screen "1002_Process Value Mixing Head" 1280x800, template "Navigation"
   on GenerateScreen: SetBit("DB704_MH_Value_Read")
   Group "Group" at 107,163 size 1065x534
   TextField "Text field_1" at 500,138 size 280x25; Text 'Process values metering unit / Process values mixing head'
   TextField "Text field_2" at 138,222 size 112x25; Text 'Module No.'
   TextField "Text field_3" at 138,256 size 81x25; Text 'Address'
   TextField "Text field_4" at 138,290 size 64x25; Text 'Offset'
   TextField "Text field_5" at 138,323 size 96x25; Text 'Multiplier'
   TextField "Text field_6" at 138,357 size 174x25; Text 'Min. Value Sensor'
   TextField "Text field_7" at 138,391 size 178x25; Text 'Max. Value Sensor'
   TextField "Text field_10" at 445,189 size 141x25; Text 'Pressure Con2'
   TextField "Text field_11" at 589,189 size 141x25; Text 'Pressure Con3'
   IOField "PV_MeteringUnit_ModulNoPressureCon1" at 313,219 size 122x30; Authorization "User administration"; FormatPattern s9999999
      ProcessValue <- "DB604_PV_Mixinghead_Mixinghead{0}_Pressure_Connection{1}_PV_Conf_ActV_ModulNo"
   IOField "I/O field_2" at 313,253 size 122x30; Authorization "User administration"; FormatPattern s9999999
      ProcessValue <- "DB604_PV_Mixinghead_Mixinghead{0}_Pressure_Connection{1}_PV_Conf_ActV_Address"
   IOField "I/O field_3" at 313,287 size 122x30; Authorization "User administration"; FormatPattern s9999999
      ProcessValue <- "DB604_PV_Mixinghead_Mixinghead{0}_Pressure_Connection{1}_PV_Conf_ActV_OffsetSignal"
   IOField "I/O field_4" at 313,321 size 122x30; Authorization "User administration"; FormatPattern s99999.999
      ProcessValue <- "DB604_PV_Mixinghead_Mixinghead{0}_Pressure_Connection{1}_PV_Conf_ActV_Multiplier"
   IOField "I/O field_5" at 313,355 size 122x30; Authorization "User administration"; FormatPattern s99999
      ProcessValue <- "DB604_PV_Mixinghead_Mixinghead{0}_Pressure_Connection{1}_PV_Conf_ActV_MinValueSensor"
   IOField "I/O field_6" at 313,389 size 122x30; Authorization "User administration"; FormatPattern s9999999
      ProcessValue <- "DB604_PV_Mixinghead_Mixinghead{0}_Pressure_Connection{1}_PV_Conf_ActV_MaxValueSensor"
   IOField "I/O field_8" at 454,219 size 122x30; Authorization "User administration"; FormatPattern s9999999
      ProcessValue <- "DB604_PV_Mixinghead_Mixinghead{0}_Pressure_Connection{2}_PV_Conf_ActV_ModulNo"
   IOField "I/O field_9" at 454,253 size 122x30; Authorization "User administration"; FormatPattern s9999999
      ProcessValue <- "DB604_PV_Mixinghead_Mixinghead{0}_Pressure_Connection{2}_PV_Conf_ActV_Address"
   IOField "I/O field_10" at 454,287 size 122x30; Authorization "User administration"; FormatPattern s9999999
      ProcessValue <- "DB604_PV_Mixinghead_Mixinghead{0}_Pressure_Connection{2}_PV_Conf_ActV_OffsetSignal"
   IOField "I/O field_11" at 454,321 size 122x30; Authorization "User administration"; FormatPattern s99999.999
      ProcessValue <- "DB604_PV_Mixinghead_Mixinghead{0}_Pressure_Connection{2}_PV_Conf_ActV_Multiplier"
   IOField "I/O field_12" at 454,355 size 122x30; Authorization "User administration"; FormatPattern s99999
      ProcessValue <- "DB604_PV_Mixinghead_Mixinghead{0}_Pressure_Connection{2}_PV_Conf_ActV_MinValueSensor"
   IOField "I/O field_13" at 454,389 size 122x30; Authorization "User administration"; FormatPattern s9999999
      ProcessValue <- "DB604_PV_Mixinghead_Mixinghead{0}_Pressure_Connection{2}_PV_Conf_ActV_MaxValueSensor"
   IOField "I/O field_14" at 598,219 size 122x30; Authorization "User administration"; FormatPattern s9999999
      ProcessValue <- "DB604_PV_Mixinghead_Mixinghead{0}_Pressure_Connection{3}_PV_Conf_ActV_ModulNo"
   IOField "I/O field_15" at 598,253 size 122x30; Authorization "User administration"; FormatPattern s9999999
      ProcessValue <- "DB604_PV_Mixinghead_Mixinghead{0}_Pressure_Connection{3}_PV_Conf_ActV_Address"
   IOField "I/O field_16" at 598,287 size 122x30; Authorization "User administration"; FormatPattern s9999999
      ProcessValue <- "DB604_PV_Mixinghead_Mixinghead{0}_Pressure_Connection{3}_PV_Conf_ActV_OffsetSignal"
   IOField "I/O field_17" at 598,321 size 122x30; Authorization "User administration"; FormatPattern s99999.999
      ProcessValue <- "DB604_PV_Mixinghead_Mixinghead{0}_Pressure_Connection{3}_PV_Conf_ActV_Multiplier"
   IOField "I/O field_18" at 598,355 size 122x30; Authorization "User administration"; FormatPattern s99999
      ProcessValue <- "DB604_PV_Mixinghead_Mixinghead{0}_Pressure_Connection{3}_PV_Conf_ActV_MinValueSensor"
   IOField "I/O field_19" at 598,389 size 122x30; Authorization "User administration"; FormatPattern s9999999
      ProcessValue <- "DB604_PV_Mixinghead_Mixinghead{0}_Pressure_Connection{3}_PV_Conf_ActV_MaxValueSensor"
   TextField "Text field_16" at 734,189 size 141x25; Text 'Pressure Con4'
   TextField "Text field_17" at 873,189 size 141x25; Text 'Pressure Con5'
   IOField "I/O field_23" at 882,219 size 122x30; Authorization "User administration"; FormatPattern s9999999
      ProcessValue <- "DB604_PV_Mixinghead_Mixinghead{0}_Pressure_Connection{5}_PV_Conf_ActV_ModulNo"
   IOField "I/O field_24" at 882,253 size 122x30; Authorization "User administration"; FormatPattern s9999999
      ProcessValue <- "DB604_PV_Mixinghead_Mixinghead{0}_Pressure_Connection{5}_PV_Conf_ActV_Address"
   IOField "I/O field_25" at 882,287 size 122x30; Authorization "User administration"; FormatPattern s9999999
      ProcessValue <- "DB604_PV_Mixinghead_Mixinghead{0}_Pressure_Connection{5}_PV_Conf_ActV_OffsetSignal"
   IOField "I/O field_26" at 882,321 size 122x30; Authorization "User administration"; FormatPattern s99999.999
      ProcessValue <- "DB604_PV_Mixinghead_Mixinghead{0}_Pressure_Connection{5}_PV_Conf_ActV_Multiplier"
   IOField "I/O field_27" at 882,355 size 122x30; Authorization "User administration"; FormatPattern s99999
      ProcessValue <- "DB604_PV_Mixinghead_Mixinghead{0}_Pressure_Connection{5}_PV_Conf_ActV_MinValueSensor"
   IOField "I/O field_28" at 882,389 size 122x30; Authorization "User administration"; FormatPattern s9999999
      ProcessValue <- "DB604_PV_Mixinghead_Mixinghead{0}_Pressure_Connection{5}_PV_Conf_ActV_MaxValueSensor"
   TextField "Text field_9" at 304,189 size 141x25; Text 'Pressure Con1'
   TextField "Text field_29" at 1014,191 size 141x25; Text 'Pressure Con6'
   IOField "I/O field_35" at 1023,219 size 122x30; Authorization "User administration"; FormatPattern s9999999
      ProcessValue <- "DB604_PV_Mixinghead_Mixinghead{0}_Pressure_Connection{6}_PV_Conf_ActV_ModulNo"
   IOField "I/O field_36" at 1023,253 size 122x30; Authorization "User administration"; FormatPattern s9999999
      ProcessValue <- "DB604_PV_Mixinghead_Mixinghead{0}_Pressure_Connection{6}_PV_Conf_ActV_Address"
   IOField "I/O field_37" at 1023,287 size 122x30; Authorization "User administration"; FormatPattern s9999999
      ProcessValue <- "DB604_PV_Mixinghead_Mixinghead{0}_Pressure_Connection{6}_PV_Conf_ActV_OffsetSignal"
   IOField "I/O field_38" at 1023,321 size 122x30; Authorization "User administration"; FormatPattern s99999.999
      ProcessValue <- "DB604_PV_Mixinghead_Mixinghead{0}_Pressure_Connection{6}_PV_Conf_ActV_Multiplier"
   IOField "I/O field_39" at 1023,355 size 122x30; Authorization "User administration"; FormatPattern s99999
      ProcessValue <- "DB604_PV_Mixinghead_Mixinghead{0}_Pressure_Connection{6}_PV_Conf_ActV_MinValueSensor"
   IOField "I/O field_40" at 1023,389 size 122x30; Authorization "User administration"; FormatPattern s9999999
      ProcessValue <- "DB604_PV_Mixinghead_Mixinghead{0}_Pressure_Connection{6}_PV_Conf_ActV_MaxValueSensor"
   IOField "I/O field_7" at 739,219 size 122x30; Authorization "User administration"; FormatPattern s9999999
      ProcessValue <- "DB604_PV_Mixinghead_Mixinghead{0}_Pressure_Connection{4}_PV_Conf_ActV_ModulNo"
   IOField "I/O field_20" at 739,253 size 122x30; Authorization "User administration"; FormatPattern s9999999
      ProcessValue <- "DB604_PV_Mixinghead_Mixinghead{0}_Pressure_Connection{4}_PV_Conf_ActV_Address"
   IOField "I/O field_21" at 739,287 size 122x30; Authorization "User administration"; FormatPattern s9999999
      ProcessValue <- "DB604_PV_Mixinghead_Mixinghead{0}_Pressure_Connection{4}_PV_Conf_ActV_OffsetSignal"
   IOField "I/O field_22" at 739,321 size 122x30; Authorization "User administration"; FormatPattern s99999.999
      ProcessValue <- "DB604_PV_Mixinghead_Mixinghead{0}_Pressure_Connection{4}_PV_Conf_ActV_Multiplier"
   IOField "I/O field_29" at 739,355 size 122x30; Authorization "User administration"; FormatPattern s99999
      ProcessValue <- "DB604_PV_Mixinghead_Mixinghead{0}_Pressure_Connection{4}_PV_Conf_ActV_MinValueSensor"
   IOField "I/O field_30" at 739,389 size 122x30; Authorization "User administration"; FormatPattern s9999999
      ProcessValue <- "DB604_PV_Mixinghead_Mixinghead{0}_Pressure_Connection{4}_PV_Conf_ActV_MaxValueSensor"
   TextField "Text field_8" at 138,462 size 112x25; Text 'Module No.'
   TextField "Text field_12" at 138,497 size 81x25; Text 'Address'
   TextField "Text field_13" at 138,532 size 64x25; Text 'Offset'
   TextField "Text field_14" at 138,566 size 96x25; Text 'Multiplier'
   TextField "Text field_15" at 138,600 size 174x25; Text 'Min. Value Sensor'
   TextField "Text field_18" at 138,634 size 178x25; Text 'Max. Value Sensor'
   TextField "Text field_19" at 460,426 size 110x25; Text 'Temp Con2'
   TextField "Text field_20" at 604,426 size 110x25; Text 'Temp Con3'
   IOField "I/O field_31" at 313,459 size 122x30; Authorization "User administration"; FormatPattern s9999999
      ProcessValue <- "DB604_PV_Mixinghead_Mixinghead{0}_Temperature_Connection{1}_PV_Conf_ActV_ModulNo"
   IOField "I/O field_32" at 313,494 size 122x30; Authorization "User administration"; FormatPattern s9999999
      ProcessValue <- "DB604_PV_Mixinghead_Mixinghead{0}_Temperature_Connection{1}_PV_Conf_ActV_Address"
   IOField "I/O field_33" at 313,529 size 122x30; Authorization "User administration"; FormatPattern s9999999
      ProcessValue <- "DB604_PV_Mixinghead_Mixinghead{0}_Temperature_Connection{1}_PV_Conf_ActV_OffsetSignal"
   IOField "I/O field_34" at 313,563 size 122x30; Authorization "User administration"; FormatPattern s99999.999
      ProcessValue <- "DB604_PV_Mixinghead_Mixinghead{0}_Temperature_Connection{1}_PV_Conf_ActV_Multiplier"
   IOField "I/O field_41" at 313,597 size 122x30; Authorization "User administration"; FormatPattern s9999999
      ProcessValue <- "DB604_PV_Mixinghead_Mixinghead{0}_Temperature_Connection{1}_PV_Conf_ActV_MinValueSensor"
   IOField "I/O field_42" at 313,631 size 122x30; Authorization "User administration"; FormatPattern s9999999
      ProcessValue <- "DB604_PV_Mixinghead_Mixinghead{0}_Temperature_Connection{1}_PV_Conf_ActV_MaxValueSensor"
   IOField "I/O field_43" at 454,458 size 122x30; Authorization "User administration"; FormatPattern s9999999
      ProcessValue <- "DB604_PV_Mixinghead_Mixinghead{0}_Temperature_Connection{2}_PV_Conf_ActV_ModulNo"
   IOField "I/O field_44" at 454,493 size 122x30; Authorization "User administration"; FormatPattern s9999999
      ProcessValue <- "DB604_PV_Mixinghead_Mixinghead{0}_Temperature_Connection{2}_PV_Conf_ActV_Address"
   IOField "I/O field_45" at 454,528 size 122x30; Authorization "User administration"; FormatPattern s9999999
      ProcessValue <- "DB604_PV_Mixinghead_Mixinghead{0}_Temperature_Connection{2}_PV_Conf_ActV_OffsetSignal"
   IOField "I/O field_46" at 454,562 size 122x30; Authorization "User administration"; FormatPattern s99999.999
      ProcessValue <- "DB604_PV_Mixinghead_Mixinghead{0}_Temperature_Connection{2}_PV_Conf_ActV_Multiplier"
   IOField "I/O field_47" at 454,596 size 122x30; Authorization "User administration"; FormatPattern s9999999
      ProcessValue <- "DB604_PV_Mixinghead_Mixinghead{0}_Temperature_Connection{2}_PV_Conf_ActV_MinValueSensor"
   IOField "I/O field_48" at 454,630 size 122x30; Authorization "User administration"; FormatPattern s9999999
      ProcessValue <- "DB604_PV_Mixinghead_Mixinghead{0}_Temperature_Connection{2}_PV_Conf_ActV_MaxValueSensor"
   IOField "I/O field_49" at 598,457 size 122x30; Authorization "User administration"; FormatPattern s9999999
      ProcessValue <- "DB604_PV_Mixinghead_Mixinghead{0}_Temperature_Connection{3}_PV_Conf_ActV_ModulNo"
   IOField "I/O field_50" at 598,492 size 122x30; Authorization "User administration"; FormatPattern s9999999
      ProcessValue <- "DB604_PV_Mixinghead_Mixinghead{0}_Temperature_Connection{3}_PV_Conf_ActV_Address"
   IOField "I/O field_51" at 598,527 size 122x30; Authorization "User administration"; FormatPattern s9999999
      ProcessValue <- "DB604_PV_Mixinghead_Mixinghead{0}_Temperature_Connection{3}_PV_Conf_ActV_OffsetSignal"
   IOField "I/O field_52" at 598,561 size 122x30; Authorization "User administration"; FormatPattern s99999.999
      ProcessValue <- "DB604_PV_Mixinghead_Mixinghead{0}_Temperature_Connection{3}_PV_Conf_ActV_Multiplier"
   IOField "I/O field_53" at 598,595 size 122x30; Authorization "User administration"; FormatPattern s9999999
      ProcessValue <- "DB604_PV_Mixinghead_Mixinghead{0}_Temperature_Connection{3}_PV_Conf_ActV_MinValueSensor"
   IOField "I/O field_54" at 598,629 size 122x30; Authorization "User administration"; FormatPattern s9999999
      ProcessValue <- "DB604_PV_Mixinghead_Mixinghead{0}_Temperature_Connection{3}_PV_Conf_ActV_MaxValueSensor"
   TextField "Text field_21" at 745,426 size 110x25; Text 'Temp Con4'
   TextField "Text field_22" at 888,426 size 110x25; Text 'Temp Con5'
   IOField "I/O field_55" at 882,460 size 122x30; Authorization "User administration"; FormatPattern s9999999
      ProcessValue <- "DB604_PV_Mixinghead_Mixinghead{0}_Temperature_Connection{5}_PV_Conf_ActV_ModulNo"
   IOField "I/O field_56" at 882,495 size 122x30; Authorization "User administration"; FormatPattern s9999999
      ProcessValue <- "DB604_PV_Mixinghead_Mixinghead{0}_Temperature_Connection{5}_PV_Conf_ActV_Address"
   IOField "I/O field_57" at 882,530 size 122x30; Authorization "User administration"; FormatPattern s9999999
      ProcessValue <- "DB604_PV_Mixinghead_Mixinghead{0}_Temperature_Connection{5}_PV_Conf_ActV_OffsetSignal"
   IOField "I/O field_58" at 882,564 size 122x30; Authorization "User administration"; FormatPattern s99999.999
      ProcessValue <- "DB604_PV_Mixinghead_Mixinghead{0}_Temperature_Connection{5}_PV_Conf_ActV_Multiplier"
   IOField "I/O field_59" at 882,598 size 122x30; Authorization "User administration"; FormatPattern s9999999
      ProcessValue <- "DB604_PV_Mixinghead_Mixinghead{0}_Temperature_Connection{5}_PV_Conf_ActV_MinValueSensor"
   IOField "I/O field_60" at 882,632 size 122x30; Authorization "User administration"; FormatPattern s9999999
      ProcessValue <- "DB604_PV_Mixinghead_Mixinghead{0}_Temperature_Connection{5}_PV_Conf_ActV_MaxValueSensor"
   TextField "Text field_23" at 319,426 size 110x25; Text 'Temp Con1'
   TextField "Text field_24" at 1029,428 size 110x25; Text 'Temp Con6'
   IOField "I/O field_61" at 1023,460 size 122x30; Authorization "User administration"; FormatPattern s9999999
      ProcessValue <- "DB604_PV_Mixinghead_Mixinghead{0}_Temperature_Connection{6}_PV_Conf_ActV_ModulNo"
   IOField "I/O field_62" at 1023,495 size 122x30; Authorization "User administration"; FormatPattern s9999999
      ProcessValue <- "DB604_PV_Mixinghead_Mixinghead{0}_Temperature_Connection{6}_PV_Conf_ActV_Address"
   IOField "I/O field_63" at 1023,530 size 122x30; Authorization "User administration"; FormatPattern s9999999
      ProcessValue <- "DB604_PV_Mixinghead_Mixinghead{0}_Temperature_Connection{6}_PV_Conf_ActV_OffsetSignal"
   IOField "I/O field_64" at 1023,564 size 122x30; Authorization "User administration"; FormatPattern s99999.999
      ProcessValue <- "DB604_PV_Mixinghead_Mixinghead{0}_Temperature_Connection{6}_PV_Conf_ActV_Multiplier"
   IOField "I/O field_65" at 1023,598 size 122x30; Authorization "User administration"; FormatPattern s9999999
      ProcessValue <- "DB604_PV_Mixinghead_Mixinghead{0}_Temperature_Connection{6}_PV_Conf_ActV_MinValueSensor"
   IOField "I/O field_66" at 1023,632 size 122x30; Authorization "User administration"; FormatPattern s9999999
      ProcessValue <- "DB604_PV_Mixinghead_Mixinghead{0}_Temperature_Connection{6}_PV_Conf_ActV_MaxValueSensor"
   IOField "I/O field_67" at 739,458 size 122x30; Authorization "User administration"; FormatPattern s9999999
      ProcessValue <- "DB604_PV_Mixinghead_Mixinghead{0}_Temperature_Connection{4}_PV_Conf_ActV_ModulNo"
   IOField "I/O field_68" at 739,493 size 122x30; Authorization "User administration"; FormatPattern s9999999
      ProcessValue <- "DB604_PV_Mixinghead_Mixinghead{0}_Temperature_Connection{4}_PV_Conf_ActV_Address"
   IOField "I/O field_69" at 739,528 size 122x30; Authorization "User administration"; FormatPattern s9999999
      ProcessValue <- "DB604_PV_Mixinghead_Mixinghead{0}_Temperature_Connection{4}_PV_Conf_ActV_OffsetSignal"
   IOField "I/O field_70" at 739,562 size 122x30; Authorization "User administration"; FormatPattern s99999.999
      ProcessValue <- "DB604_PV_Mixinghead_Mixinghead{0}_Temperature_Connection{4}_PV_Conf_ActV_Multiplier"
   IOField "I/O field_71" at 739,596 size 122x30; Authorization "User administration"; FormatPattern s9999999
      ProcessValue <- "DB604_PV_Mixinghead_Mixinghead{0}_Temperature_Connection{4}_PV_Conf_ActV_MinValueSensor"
   IOField "I/O field_72" at 739,630 size 122x30; Authorization "User administration"; FormatPattern s9999999
      ProcessValue <- "DB604_PV_Mixinghead_Mixinghead{0}_Temperature_Connection{4}_PV_Conf_ActV_MaxValueSensor"
   TextField "Text field_25" at 266,706 size 81x25; Text 'Address'
   TextField "Text field_26" at 266,736 size 64x25; Text 'Offset'
   TextField "Text field_27" at 266,764 size 96x25; Text 'Multiplier'
   TextField "Text field_28" at 418,706 size 371x25; Text 'Address Number PLC or ProCan Chanel'
   TextField "Text field_30" at 418,736 size 321x25; Text 'Value to add the calculated value'
   TextField "Text field_31" at 418,764 size 659x25; Text 'conversion value for the actual value (signal detail/max.value x100)'
   SymbolicIOField "Symbolic I/O field_1" at 326,104 size 451x32; TextOn '1'; TextOff '0'; TextList "MH_IOField"
      ProcessValue <- "DB614_MH_State_ReadDeviceNo"
   Button "b_Incress_PV_MeteringUnit" at 788,104 size 46x32; TextOff 'Text'; PictureOff "NEXT"
      on Press: function_dd21b452("DB614_MH_State_ReadDeviceNo", 1)
   Button "b_Decress_PV_MeteringUnit" at 270,104 size 46x32; TextOff 'Text'; PictureOff "BEFORE"
      on Press: function_b9b71300("DB614_MH_State_ReadDeviceNo", 1)

screen "1005_Process Value MH Inerting" 1280x800, template "Navigation"
   on GenerateScreen: SetBit("DB704_MH_Value_Read")
   Group "Group" at 118,178 size 672x493
   TextField "Text field_2" at 243,258 size 112x25; Text 'Module No.'
   TextField "Text field_3" at 243,306 size 81x25; Text 'Address'
   TextField "Text field_4" at 243,354 size 64x25; Text 'Offset'
   TextField "Text field_5" at 243,402 size 96x25; Text 'Multiplier'
   TextField "Text field_6" at 243,450 size 174x25; Text 'Min. Value Sensor'
   TextField "Text field_7" at 243,498 size 178x25; Text 'Max. Value Sensor'
   TextField "Text field_8" at 243,606 size 123x25; Text 'Actual Value'
   TextField "Text field_9" at 511,208 size 83x25; Text 'Inerting'
   IOField "PV_inerting_ModuleNo" at 481,255 size 142x30; Authorization "User administration"; FormatPattern 9999999
      ProcessValue <- "DB604_PV_Mixinghead_Mixinghead{0}_Inerting_PV_Conf_ActV_ModulNo"
   IOField "I/O field_2" at 481,303 size 142x30; Authorization "User administration"; FormatPattern 9999999
      ProcessValue <- "DB604_PV_Mixinghead_Mixinghead{0}_Inerting_PV_Conf_ActV_Address"
   IOField "I/O field_3" at 481,351 size 142x30; Authorization "User administration"; FormatPattern 9999999
      ProcessValue <- "DB604_PV_Mixinghead_Mixinghead{0}_Inerting_PV_Conf_ActV_OffsetSignal"
   IOField "I/O field_4" at 481,399 size 142x30; Authorization "User administration"; FormatPattern 99999.999
      ProcessValue <- "DB604_PV_Mixinghead_Mixinghead{0}_Inerting_PV_Conf_ActV_Multiplier"
   IOField "I/O field_5" at 481,447 size 142x30; Authorization "User administration"; FormatPattern 9999999
      ProcessValue <- "DB604_PV_Mixinghead_Mixinghead{0}_Inerting_PV_Conf_ActV_MinValueSensor"
   IOField "I/O field_6" at 481,495 size 142x30; Authorization "User administration"; FormatPattern 9999999
      ProcessValue <- "DB604_PV_Mixinghead_Mixinghead{0}_Inerting_PV_Conf_ActV_MaxValueSensor"
   IOField "I/O field_7" at 481,603 size 142x30; Authorization "User administration"; FormatPattern 9999999
      ProcessValue <- "DB604_PV_Mixinghead_Mixinghead{0}_Inerting_PV_ActV_Value"
   SymbolicIOField "Symbolic I/O field_1" at 326,104 size 451x32; TextOn '1'; TextOff '0'; TextList "MH_IOField"
      ProcessValue <- "DB614_MH_State_ReadDeviceNo"
   TextField "Text field_10" at 505,552 size 94x25; Text '[NL/min]'
   Button "b_Incress_PV_Inerting" at 787,104 size 46x32; TextOff 'Text'; PictureOff "NEXT"
      on Click: function_dd21b452("DB614_MH_State_ReadDeviceNo", 1)
   Button "b_Decress_PV_inerting" at 272,104 size 46x32; TextOff 'Text'; PictureOff "BEFORE"
      on Click: function_b9b71300("DB614_MH_State_ReadDeviceNo", 1)

screen "2004_ProNet MH digital" 1280x800, template "Navigation"
   on GenerateScreen: SetBit("PN_Mixinghead_Send"); SetBit("PN_Mixinghead_Mixinghead{0}_Digital_GeneralParameters_Request")
   Group "Group" at 118,180 size 1041x561
   TextField "Text field_1" at 428,143 size 247x29; Text 'ProNet Configuration'
   TextField "Text field_3" at 290,258 size 122x25; Text 'Start Adress'
   TextField "Text field_4" at 291,308 size 186x25; Text 'MixingHead Chanel'
   TextField "Text field_5" at 292,358 size 320x25; Text 'MixingHead valve output number'
   TextField "Text field_6" at 293,408 size 413x25; Text 'Mixinghead proximity switch input number'
   TextField "Text field_7" at 294,458 size 408x25; Text 'MixingHead external release input number'
   TextField "Text field_8" at 295,508 size 332x25; Text 'Monitoring time mixing head open'
   TextField "Text field_9" at 296,558 size 334x25; Text 'Monitoring time mixing head close'
   TextField "Text field_10" at 297,608 size 223x25; Text 'Allowed bouncing time'
   TextField "Text field_11" at 298,658 size 298x25; Text 'Delay time for external release'
   TextField "Text field_12" at 860,658 size 46x25; Text '[s]'
   TextField "Text field_13" at 860,608 size 46x25; Text '[s]'
   TextField "Text field_14" at 860,558 size 46x25; Text '[s]'
   TextField "Text field_15" at 860,508 size 46x25; Text '[s]'
   IOField "Monitoring_Time _Mixinghead_Open" at 752,505 size 96x32; FormatPattern 999999.999
      ProcessValue <- "PN_Mixinghead_Mixinghead{0}_Digital_Zeiten_Data_ÜberwachungszeitÖffnen"
   IOField "I/O field_2" at 752,555 size 96x32; FormatPattern 999999.999
      ProcessValue <- "PN_Mixinghead_Mixinghead{0}_Digital_Zeiten_Data_ÜberwachungszeitSchließen"
   IOField "I/O field_3" at 752,605 size 96x32; FormatPattern 999999.999
      ProcessValue <- "PN_Mixinghead_Mixinghead{0}_Digital_Zeiten_Data_ErlaubtePrellzeit"
   IOField "I/O field_4" at 752,255 size 96x32; FormatPattern 99999
      ProcessValue <- "PN_Mixinghead_Mixinghead{0}_Digital_Address"
   Button "Button_1" at 872,253 size 96x32; TextOff 'Active'
      on Press: InvertBit("PN_Mixinghead_Mixinghead{0}_Digital_Active"); SetBit("PN_Mixinghead_Mixinghead{0}_Digital_GeneralParameters_Request"); SetBit("PN_Mixinghead_Mixinghead{0}_Digital_Zeiten_2_Request"); SetBit("PN_Mixinghead_Mixinghead{0}_Digital_Zeiten_Request")
      Appearance <- "PN_Mixinghead_Mixinghead{0}_Digital_Active"
   SymbolicIOField "Symbolic I/O field_1" at 752,296 size 96x32; TextOff '0'; TextOn '1'; TextList "Pronet_Mixinghead Chanel"
      ProcessValue <- "PN_Mixinghead_Mixinghead{0}_Digital_GeneralParameters_Data_MischkopfKanal"
   SymbolicIOField "Symbolic I/O field_2" at 752,344 size 96x32; TextOn '1'; TextOff '0'; TextList "Pronet_Mixinghead_Output_Valve_Numb"
      ProcessValue <- "PN_Mixinghead_Mixinghead{0}_Digital_GeneralParameters_Data_Ventilausgang"
   SymbolicIOField "Symbolic I/O field_3" at 752,400 size 96x32; TextOn '1'; TextOff '0'; TextList "Pronet_Proximity_switch_Input"
      ProcessValue <- "PN_Mixinghead_Mixinghead{0}_Digital_GeneralParameters_Data_EingangskanalMK_Ini"
   SymbolicIOField "Symbolic I/O field_4" at 752,453 size 96x32; TextOn '1'; TextOff '0'; TextList "Pronet_External_Release_Switch_Input"
      ProcessValue <- "PN_Mixinghead_Mixinghead{0}_Digital_GeneralParameters_Data_EingangskanalFreigabe"
   IOField "I/O field_5" at 752,656 size 96x32; FormatPattern 999999.999
      ProcessValue <- "PN_Mixinghead_Mixinghead{0}_Digital_Zeiten_2_Data_Verzögerungszeit_HW_Freigabe"
   SymbolicIOField "Symbolic I/O field_5" at 326,104 size 451x32; TextOff '0'; TextOn '1'; TextList "MH_NO"
      ProcessValue <- "PN_Mixinghead_SetIndex"
   Button "b_Incress_Pronet_Mixinghead" at 787,104 size 46x32; TextOff 'Text'; PictureOff "NEXT"
      on Press: function_dd21b452("PN_Mixinghead_SetIndex", 1); SetBit("PN_Mixinghead_Send")
   Button "b_Decress_Pronet_Mixinghead" at 270,104 size 46x32; TextOff 'Text'; PictureOff "BEFORE"
      on Press: function_b9b71300("PN_Mixinghead_SetIndex", 1); SetBit("PN_Mixinghead_Send")
   TextField "Text field_2" at 438,207 size 227x29; Text 'Mixinghead Control'

screen "2003_ProNet CP digital" 1280x800, template "Navigation"
   on GenerateScreen: SetBit("PN_Mixinghead_Send")
   Group "Group" at 118,194 size 1041x564
   TextField "Text field_3" at 280,293 size 122x25; Text 'Start Adress'
   TextField "Text field_4" at 280,333 size 198x25; Text 'MixingHead Channel'
   TextField "Text field_5" at 280,373 size 357x25; Text 'Cleaning piston valve output number'
   TextField "Text field_6" at 280,413 size 386x25; Text 'Cleaning proximity switch input number'
   TextField "Text field_7" at 280,518 size 304x25; Text 'Monitoring time piston forward'
   TextField "Text field_8" at 280,558 size 320x25; Text 'Monitoring time piston backward'
   TextField "Text field_9" at 280,598 size 223x25; Text 'Allowed bouncing time'
   TextField "Text field_10" at 280,638 size 315x25; Text 'Waiting time in forward position'
   TextField "Text field_11" at 280,678 size 299x25; Text 'Delay time for request forward'
   TextField "Text field_12" at 906,678 size 46x25; Text '[s]'
   TextField "Text field_13" at 906,638 size 46x25; Text '[s]'
   TextField "Text field_14" at 906,598 size 46x25; Text '[s]'
   TextField "Text field_15" at 906,558 size 46x25; Text '[s]'
   TextField "Text field_16" at 906,518 size 46x25; Text '[s]'
   SymbolicIOField "Symbolic I/O field_5" at 326,104 size 451x32; TextOn '1'; TextOff '0'; TextList "MH_NO"
      ProcessValue <- "PN_Mixinghead_SetIndex"
   Button "b_Incress_CleaningPiston_Control" at 787,104 size 46x32; TextOff 'Text'; PictureOff "NEXT"
      on Press: function_dd21b452("PN_Mixinghead_SetIndex", 1); SetBit("PN_Mixinghead_Send")
   Button "b_Decress_CleaningPiston_Control" at 270,104 size 46x32; TextOff 'Text'; PictureOff "BEFORE"
      on Press: function_b9b71300("PN_Mixinghead_SetIndex", 1); SetBit("PN_Mixinghead_Send")
   TextField "Text field_1" at 428,147 size 247x29; Text 'ProNet Configuration'
   IOField "Start_Adress_Cleaning Piston Control" at 808,290 size 96x32; FormatPattern 999999
      ProcessValue <- "PN_Mixinghead_Mixinghead{0}_ReinigungskolbenDigital_Address"
   Button "Button_1" at 928,290 size 96x32; TextOff 'Active'
      on Press: InvertBit("PN_Mixinghead_Mixinghead{0}_ReinigungskolbenDigital_Active")
      Appearance <- "PN_Mixinghead_Mixinghead{0}_ReinigungskolbenDigital_Active"
   IOField "I/O field_2" at 808,515 size 96x32; FormatPattern 99999.999
      ProcessValue <- "PN_Mixinghead_Mixinghead{0}_ReinigungskolbenDigital_Zeiten_Data_ÜberwachungszeitVorfahren"
   IOField "I/O field_3" at 808,555 size 96x32; FormatPattern 99999.999
      ProcessValue <- "PN_Mixinghead_Mixinghead{0}_ReinigungskolbenDigital_Zeiten_Data_ÜberwachungszeitRückfahren"
   IOField "I/O field_4" at 808,595 size 96x32; FormatPattern 99999.999
      ProcessValue <- "PN_Mixinghead_Mixinghead{0}_ReinigungskolbenDigital_Zeiten_Data_ErlaubtePrellzeit"
   SymbolicIOField "Symbolic I/O field_1" at 808,330 size 96x32; TextOn '1'; TextOff '0'; TextList "Pronet_Mixinghead Chanel"
      ProcessValue <- "PN_Mixinghead_Mixinghead{0}_ReinigungskolbenDigital_GeneralParameters_Data_MischkopfKanal"
   SymbolicIOField "Symbolic I/O field_2" at 808,370 size 96x32; TextOn '1'; TextOff '0'; TextList "Pronet_Mixinghead_Output_Valve_Numb"
      ProcessValue <- "PN_Mixinghead_Mixinghead{0}_ReinigungskolbenDigital_GeneralParameters_Data_AusgangRKVentil"
   SymbolicIOField "Symbolic I/O field_3" at 808,410 size 96x32; TextOn '1'; TextOff '0'; TextList "Pronet_Proximity_switch_Input"
      ProcessValue <- "PN_Mixinghead_Mixinghead{0}_ReinigungskolbenDigital_GeneralParameters_Data_EingangskanalRK_Ini"
   IOField "I/O field_5" at 808,675 size 96x32; FormatPattern 99999.999
      ProcessValue <- "PN_Mixinghead_Mixinghead{0}_ReinigungskolbenDigital_Zeiten_Data_VerzögerungNachSchuss"
   IOField "I/O field_6" at 808,635 size 96x32; FormatPattern 99999.999
      ProcessValue <- "PN_Mixinghead_Mixinghead{0}_ReinigungskolbenDigital_Zeiten_Data_WartezeitVorne"
   TextField "Text field_2" at 415,224 size 273x29; Text 'Cleaning Piston Control'

screen "2001_ProNet analog input" 1280x800, template "Navigation"
   Group "Group" at 118,225 size 1041x545
   TextField "Text field_3" at 170,348 size 56x25; Text 'Mode'
   TextField "Text field_4" at 170,388 size 172x25; Text 'Volltage_ZeroPos'
   TextField "Text field_5" at 170,430 size 105x25; Text 'Value_10V'
   TextField "Text field_6" at 170,470 size 139x25; Text 'Tank_Average'
   TextField "Text field_7" at 457,573 size 254x25; Text '0:0.. 5 V; 1: -5.. +5 V;'
   TextField "Text field_8" at 690,573 size 308x25; Text '2:0.. 10 V; 3: -10 V.. +10 V;'
   TextField "Text field_9" at 222,573 size 56x25; Text 'Mode'
   TextField "Text field_10" at 222,613 size 172x25; Text 'Volltage_ZeroPos'
   TextField "Text field_11" at 222,652 size 105x25; Text 'Value_10V'
   TextField "Text field_12" at 222,692 size 139x25; Text 'Tank_Average'
   TextField "Text field_13" at 458,612 size 578x25; Text 'Voltage [mV] at min. input value (if 4...20mA 2000 inscribe)'
   TextField "Text field_14" at 457,652 size 366x25; Text 'Max Value for input 10V or 138.5 ohm'
   TextField "Text field_15" at 456,692 size 222x25; Text 'Time for average [ms]'
   TextField "Text field_16" at 371,302 size 17x25; Text '1'
   TextField "Text field_17" at 467,302 size 46x25; Text '2'
   TextField "Text field_18" at 563,302 size 46x25; Text '3'
   TextField "Text field_19" at 659,302 size 46x25; Text '4'
   TextField "Text field_20" at 755,302 size 46x25; Text '5'
   TextField "Text field_21" at 851,302 size 46x25; Text '6'
   TextField "Text field_22" at 947,302 size 46x25; Text '7'
   TextField "Text field_23" at 1043,302 size 46x25; Text '8'
   SymbolicIOField "Symbolic I/O field_5" at 326,104 size 451x32; TextOn '1'; TextOff '0'; TextList "Pronet_Analog_Input"
      ProcessValue <- "PN_AI_SetIndex"
   Button "b_Incress_AI_Control" at 786,104 size 46x32; TextOff 'Text'; PictureOff "NEXT"
      on Press: function_dd21b452("PN_AI_SetIndex", 1)
   Button "b_Decress_AI_Control" at 269,104 size 46x32; TextOff 'Text'; PictureOff "BEFORE"
      on Press: function_b9b71300("PN_AI_SetIndex", 1)
   Button "Button_1" at 1016,139 size 96x32; TextOff 'Active'
      on Press: InvertBit("PN_AI_Module{0}_AI8_Active")
      Appearance <- "PN_AI_Module{0}_AI8_Active"
   TextField "Text field_1" at 428,145 size 247x29; Text 'ProNet Configuration'
   IOField "PronetModeAI_Control_IOField" at 339,344 size 80x32; FormatPattern 9
      ProcessValue <- "PN_AI_Module{0}_AI8_X14_0_Data_Data[1]_Betriebsart"
   IOField "I/O field_2" at 435,344 size 80x32; FormatPattern 9
      ProcessValue <- "PN_AI_Module{0}_AI8_X14_0_Data_Data[2]_Betriebsart"
   IOField "I/O field_3" at 531,344 size 80x32; FormatPattern 9
      ProcessValue <- "PN_AI_Module{0}_AI8_X14_0_Data_Data[3]_Betriebsart"
   IOField "I/O field_4" at 627,344 size 80x32; FormatPattern 9
      ProcessValue <- "PN_AI_Module{0}_AI8_X14_0_Data_Data[4]_Betriebsart"
   IOField "I/O field_5" at 723,344 size 80x32; FormatPattern 9
      ProcessValue <- "PN_AI_Module{0}_AI8_X14_0_Data_Data[5]_Betriebsart"
   IOField "I/O field_6" at 819,344 size 80x32; FormatPattern 9
      ProcessValue <- "PN_AI_Module{0}_AI8_X14_0_Data_Data[6]_Betriebsart"
   IOField "I/O field_7" at 915,344 size 80x32; FormatPattern 9
      ProcessValue <- "PN_AI_Module{0}_AI8_X14_0_Data_Data[7]_Betriebsart"
   IOField "I/O field_8" at 1011,344 size 80x32; FormatPattern 9
      ProcessValue <- "PN_AI_Module{0}_AI8_X14_0_Data_Data[8]_Betriebsart"
   IOField "I/O field_9" at 339,384 size 80x32; FormatPattern s9999999
      ProcessValue <- "PN_AI_Module{0}_AI8_X14_0_Data_Data[1]_Bereichsuntergrenze"
   IOField "I/O field_10" at 435,384 size 80x32; FormatPattern s9999999
      ProcessValue <- "PN_AI_Module{0}_AI8_X14_0_Data_Data[2]_Bereichsuntergrenze"
   IOField "I/O field_11" at 531,384 size 80x32; FormatPattern s9999999
      ProcessValue <- "PN_AI_Module{0}_AI8_X14_0_Data_Data[3]_Bereichsuntergrenze"
   IOField "I/O field_12" at 627,384 size 80x32; FormatPattern s9999999
      ProcessValue <- "PN_AI_Module{0}_AI8_X14_0_Data_Data[4]_Bereichsuntergrenze"
   IOField "I/O field_13" at 723,384 size 80x32; FormatPattern s9999999
      ProcessValue <- "PN_AI_Module{0}_AI8_X14_0_Data_Data[5]_Bereichsuntergrenze"
   IOField "I/O field_14" at 819,384 size 80x32; FormatPattern s9999999
      ProcessValue <- "PN_AI_Module{0}_AI8_X14_0_Data_Data[6]_Bereichsuntergrenze"
   IOField "I/O field_15" at 915,384 size 80x32; FormatPattern s9999999
      ProcessValue <- "PN_AI_Module{0}_AI8_X14_0_Data_Data[7]_Bereichsuntergrenze"
   IOField "I/O field_16" at 1011,384 size 80x32; FormatPattern s9999999
      ProcessValue <- "PN_AI_Module{0}_AI8_X14_0_Data_Data[8]_Bereichsuntergrenze"
   IOField "I/O field_17" at 339,426 size 80x32; FormatPattern 9999
      ProcessValue <- "PN_AI_Module{0}_AI8_X14_0_Data_Data[1]_Bereichsobergrenze"
   IOField "I/O field_18" at 435,426 size 80x32; FormatPattern 9999
      ProcessValue <- "PN_AI_Module{0}_AI8_X14_0_Data_Data[2]_Bereichsobergrenze"
   IOField "I/O field_19" at 531,426 size 80x32; FormatPattern 9999
      ProcessValue <- "PN_AI_Module{0}_AI8_X14_0_Data_Data[3]_Bereichsobergrenze"
   IOField "I/O field_20" at 627,426 size 80x32; FormatPattern 9999
      ProcessValue <- "PN_AI_Module{0}_AI8_X14_0_Data_Data[4]_Bereichsobergrenze"
   IOField "I/O field_21" at 723,426 size 80x32; FormatPattern 9999
      ProcessValue <- "PN_AI_Module{0}_AI8_X14_0_Data_Data[5]_Bereichsobergrenze"
   IOField "I/O field_22" at 819,426 size 80x32; FormatPattern 9999
      ProcessValue <- "PN_AI_Module{0}_AI8_X14_0_Data_Data[6]_Bereichsobergrenze"
   IOField "I/O field_23" at 915,426 size 80x32; FormatPattern 9999
      ProcessValue <- "PN_AI_Module{0}_AI8_X14_0_Data_Data[7]_Bereichsobergrenze"
   IOField "I/O field_24" at 1011,426 size 80x32; FormatPattern 9999
      ProcessValue <- "PN_AI_Module{0}_AI8_X14_0_Data_Data[8]_Bereichsobergrenze"
   IOField "I/O field_25" at 339,466 size 80x32; FormatPattern 9999
      ProcessValue <- "PN_AI_Module{0}_AI8_X14_0_Data_Data[1]_Mittelwertzeit"
   IOField "I/O field_26" at 435,466 size 80x32; FormatPattern 9999
      ProcessValue <- "PN_AI_Module{0}_AI8_X14_0_Data_Data[2]_Mittelwertzeit"
   IOField "I/O field_27" at 531,466 size 80x32; FormatPattern 9999
      ProcessValue <- "PN_AI_Module{0}_AI8_X14_0_Data_Data[3]_Mittelwertzeit"
   IOField "I/O field_28" at 627,466 size 80x32; FormatPattern 9999
      ProcessValue <- "PN_AI_Module{0}_AI8_X14_0_Data_Data[4]_Mittelwertzeit"
   IOField "I/O field_29" at 723,466 size 80x32; FormatPattern 9999
      ProcessValue <- "PN_AI_Module{0}_AI8_X14_0_Data_Data[5]_Mittelwertzeit"
   IOField "I/O field_30" at 819,466 size 80x32; FormatPattern 9999
      ProcessValue <- "PN_AI_Module{0}_AI8_X14_0_Data_Data[6]_Mittelwertzeit"
   IOField "I/O field_31" at 915,466 size 80x32; FormatPattern 9999
      ProcessValue <- "PN_AI_Module{0}_AI8_X14_0_Data_Data[7]_Mittelwertzeit"
   IOField "I/O field_32" at 1011,466 size 80x32; FormatPattern 9999
      ProcessValue <- "PN_AI_Module{0}_AI8_X14_0_Data_Data[8]_Mittelwertzeit"
   IOField "I/O field_33" at 1016,181 size 96x32; FormatPattern 99999
      ProcessValue <- "PN_AI_Module{0}_AI8_Address"
   TextField "Text field_2" at 887,184 size 122x25; Text 'Start Adress'
   TextField "Text field_24" at 652,265 size 149x29; Text 'Analog input'